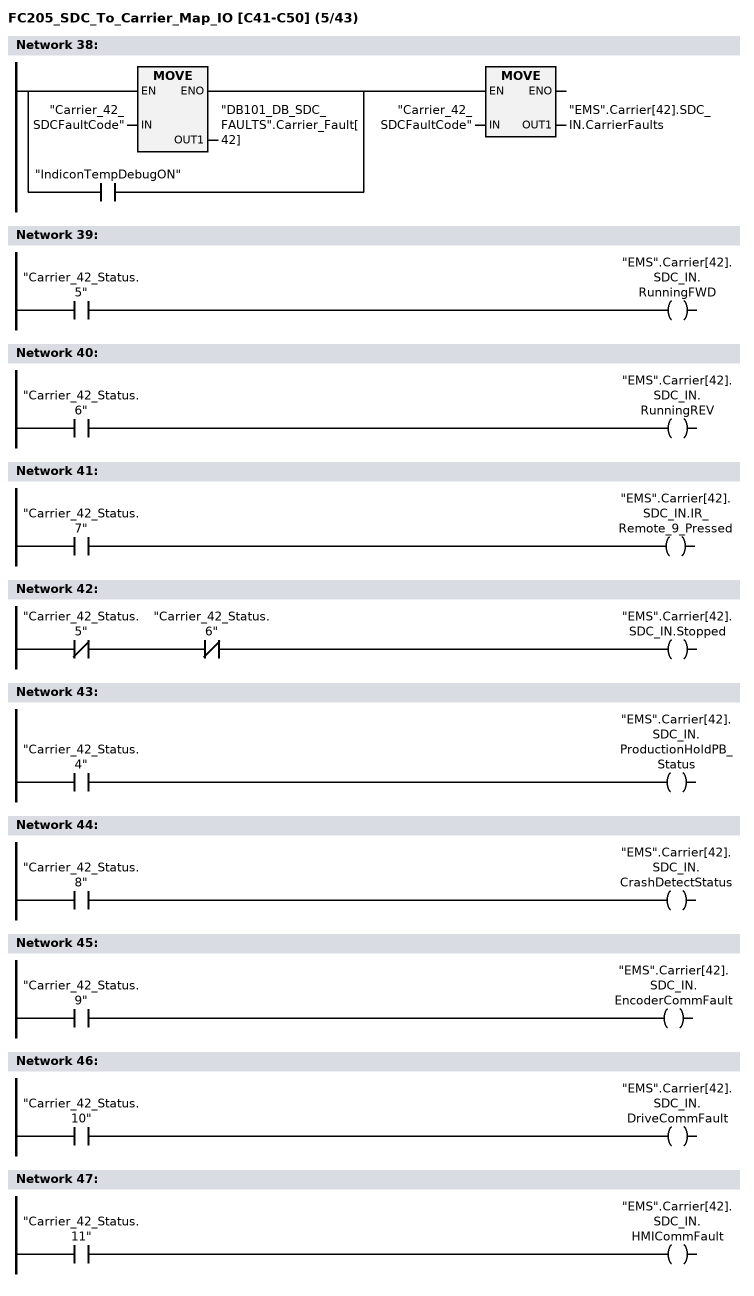
   RUNG wire#powerrail
      Move(in := "Carrier_42_SDCFaultCode", out1 => "DB101_DB_SDC_FAULTS".Carrier_Fault[42])
      wire#w1
      Move(in := "Carrier_42_SDCFaultCode", out1 => "EMS".Carrier[42].SDC_IN.CarrierFaults)
   END_RUNG
   RUNG wire#powerrail
      Contact( "IndiconTempDebugON" )
   END_RUNG wire#w1
   // the same network as SCL:
   "DB101_DB_SDC_FAULTS".Carrier_Fault[42] := "Carrier_42_SDCFaultCode";
   IF TRUE OR "IndiconTempDebugON" THEN
       "EMS".Carrier[42].SDC_IN.CarrierFaults := "Carrier_42_SDCFaultCode";
   END_IF;
END_REGION

REGION Network 39
   RUNG wire#powerrail
      Contact( "Carrier_42_Status.5" )
      Coil( "EMS".Carrier[42].SDC_IN.RunningFWD )
   END_RUNG
   // the same network as SCL:
   "EMS".Carrier[42].SDC_IN.RunningFWD := "Carrier_42_Status.5";
END_REGION

REGION Network 40
   RUNG wire#powerrail
      Contact( "Carrier_42_Status.6" )
      Coil( "EMS".Carrier[42].SDC_IN.RunningREV )
   END_RUNG
   // the same network as SCL:
   "EMS".Carrier[42].SDC_IN.RunningREV := "Carrier_42_Status.6";
END_REGION

REGION Network 41
   RUNG wire#powerrail
      Contact( "Carrier_42_Status.7" )
      Coil( "EMS".Carrier[42].SDC_IN.IR_Remote_9_Pressed )
   END_RUNG
   // the same network as SCL:
   "EMS".Carrier[42].SDC_IN.IR_Remote_9_Pressed := "Carrier_42_Status.7";
END_REGION

REGION Network 42
   RUNG wire#powerrail
      I_Contact( "Carrier_42_Status.5" )
      I_Contact( "Carrier_42_Status.6" )
      Coil( "EMS".Carrier[42].SDC_IN.Stopped )
   END_RUNG
   // the same network as SCL:
   "EMS".Carrier[42].SDC_IN.Stopped := NOT "Carrier_42_Status.5" AND NOT "Carrier_42_Status.6";
END_REGION

REGION Network 43
   RUNG wire#powerrail
      Contact( "Carrier_42_Status.4" )
      Coil( "EMS".Carrier[42].SDC_IN.ProductionHoldPB_Status )
   END_RUNG
   // the same network as SCL:
   "EMS".Carrier[42].SDC_IN.ProductionHoldPB_Status := "Carrier_42_Status.4";
END_REGION

REGION Network 44
   RUNG wire#powerrail
      Contact( "Carrier_42_Status.8" )
      Coil( "EMS".Carrier[42].SDC_IN.CrashDetectStatus )
   END_RUNG
   // the same network as SCL:
   "EMS".Carrier[42].SDC_IN.CrashDetectStatus := "Carrier_42_Status.8";
END_REGION

REGION Network 45
   RUNG wire#powerrail
      Contact( "Carrier_42_Status.9" )
      Coil( "EMS".Carrier[42].SDC_IN.EncoderCommFault )
   END_RUNG
   // the same network as SCL:
   "EMS".Carrier[42].SDC_IN.EncoderCommFault := "Carrier_42_Status.9";
END_REGION

REGION Network 46
   RUNG wire#powerrail
      Contact( "Carrier_42_Status.10" )
      Coil( "EMS".Carrier[42].SDC_IN.DriveCommFault )
   END_RUNG
   // the same network as SCL:
   "EMS".Carrier[42].SDC_IN.DriveCommFault := "Carrier_42_Status.10";
END_REGION

REGION Network 47
   RUNG wire#powerrail
      Contact( "Carrier_42_Status.11" )
      Coil( "EMS".Carrier[42].SDC_IN.HMICommFault )
   END_RUNG
   // the same network as SCL:
   "EMS".Carrier[42].SDC_IN.HMICommFault := "Carrier_42_Status.11";
END_REGION

REGION Network 48
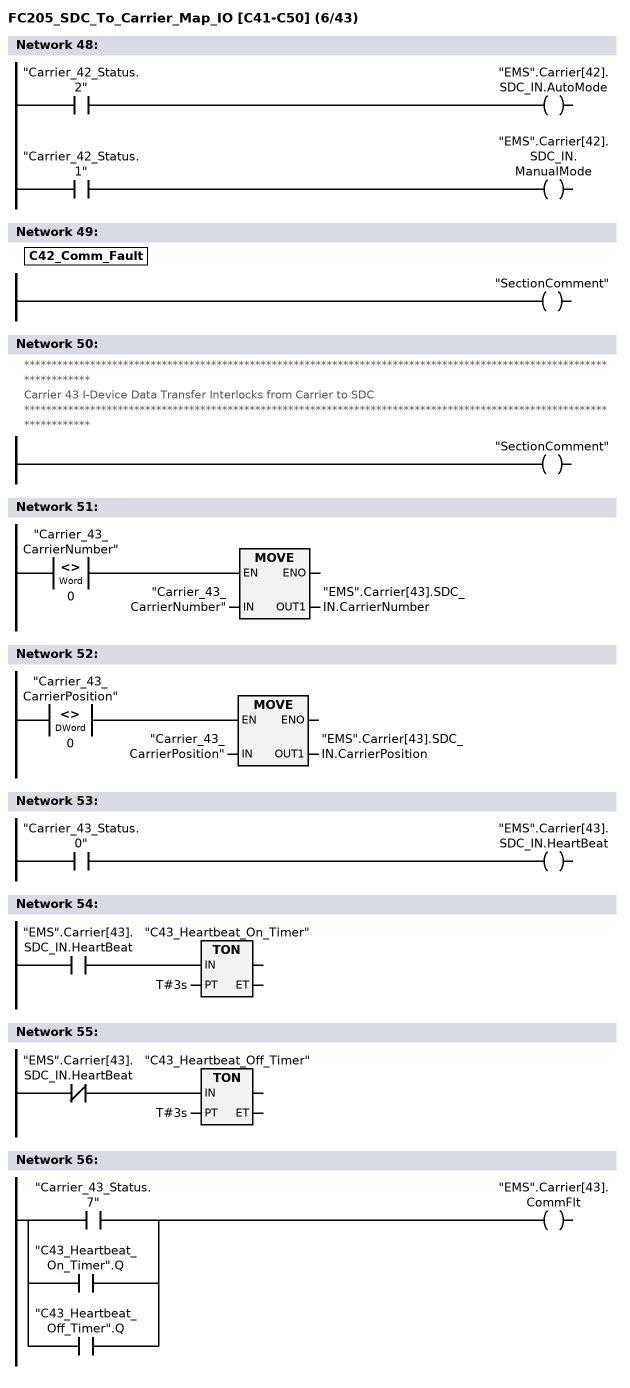
   RUNG wire#powerrail
      Contact( "Carrier_42_Status.2" )
      Coil( "EMS".Carrier[42].SDC_IN.AutoMode )
   END_RUNG
   RUNG wire#powerrail
      Contact( "Carrier_42_Status.1" )
      Coil( "EMS".Carrier[42].SDC_IN.ManualMode )
   END_RUNG
   // the same network as SCL:
   "EMS".Carrier[42].SDC_IN.AutoMode := "Carrier_42_Status.2";
   "EMS".Carrier[42].SDC_IN.ManualMode := "Carrier_42_Status.1";
END_REGION

REGION Network 49
   Label( C42_Comm_Fault )
   RUNG wire#powerrail
      Coil( "SectionComment" )
   END_RUNG
   // the same network as SCL:
   C42_Comm_Fault:
   "SectionComment" := TRUE;
END_REGION

REGION Network 50
   // **********************************************************************************************************************
   // 
   // Carrier 43 I-Device Data Transfer Interlocks from Carrier to SDC
   // 
   // **********************************************************************************************************************
   RUNG wire#powerrail
      Coil( "SectionComment" )
   END_RUNG
   // the same network as SCL:
   "SectionComment" := TRUE;
END_REGION

REGION Network 51
   RUNG wire#powerrail
      { S7_Templates := "SrcType := Word" } NE_Contact(in1 := "Carrier_43_CarrierNumber", in2 := 0)
      Move(in := "Carrier_43_CarrierNumber", out1 => "EMS".Carrier[43].SDC_IN.CarrierNumber)
   END_RUNG
   // the same network as SCL:
   IF "Carrier_43_CarrierNumber" <> 0 THEN
       "EMS".Carrier[43].SDC_IN.CarrierNumber := "Carrier_43_CarrierNumber";
   END_IF;
END_REGION

REGION Network 52
   RUNG wire#powerrail
      { S7_Templates := "SrcType := DWord" } NE_Contact(in1 := "Carrier_43_CarrierPosition", in2 := 0)
      Move(in := "Carrier_43_CarrierPosition", out1 => "EMS".Carrier[43].SDC_IN.CarrierPosition)
   END_RUNG
   // the same network as SCL:
   IF "Carrier_43_CarrierPosition" <> 0 THEN
       "EMS".Carrier[43].SDC_IN.CarrierPosition := "Carrier_43_CarrierPosition";
   END_IF;
END_REGION

REGION Network 53
   RUNG wire#powerrail
      Contact( "Carrier_43_Status.0" )
      Coil( "EMS".Carrier[43].SDC_IN.HeartBeat )
   END_RUNG
   // the same network as SCL:
   "EMS".Carrier[43].SDC_IN.HeartBeat := "Carrier_43_Status.0";
END_REGION

REGION Network 54
   "C43_Heartbeat_On_Timer".TON(IN := "EMS".Carrier[43].SDC_IN.HeartBeat, PT := T#3s);
END_REGION

REGION Network 55
   "C43_Heartbeat_Off_Timer".TON(IN := NOT "EMS".Carrier[43].SDC_IN.HeartBeat, PT := T#3s);
END_REGION

REGION Network 56
   RUNG wire#powerrail
      Contact( "Carrier_43_Status.7" )
      wire#w1
      Coil( "EMS".Carrier[43].CommFlt )
   END_RUNG
   RUNG wire#powerrail
      Contact( "C43_Heartbeat_On_Timer".Q )
   END_RUNG wire#w1
   RUNG wire#powerrail
      Contact( "C43_Heartbeat_Off_Timer".Q )
   END_RUNG wire#w1
   // the same network as SCL:
   "EMS".Carrier[43].CommFlt := "Carrier_43_Status.7" OR "C43_Heartbeat_On_Timer".Q OR "C43_Heartbeat_Off_Timer".Q;
END_REGION

REGION Network 57
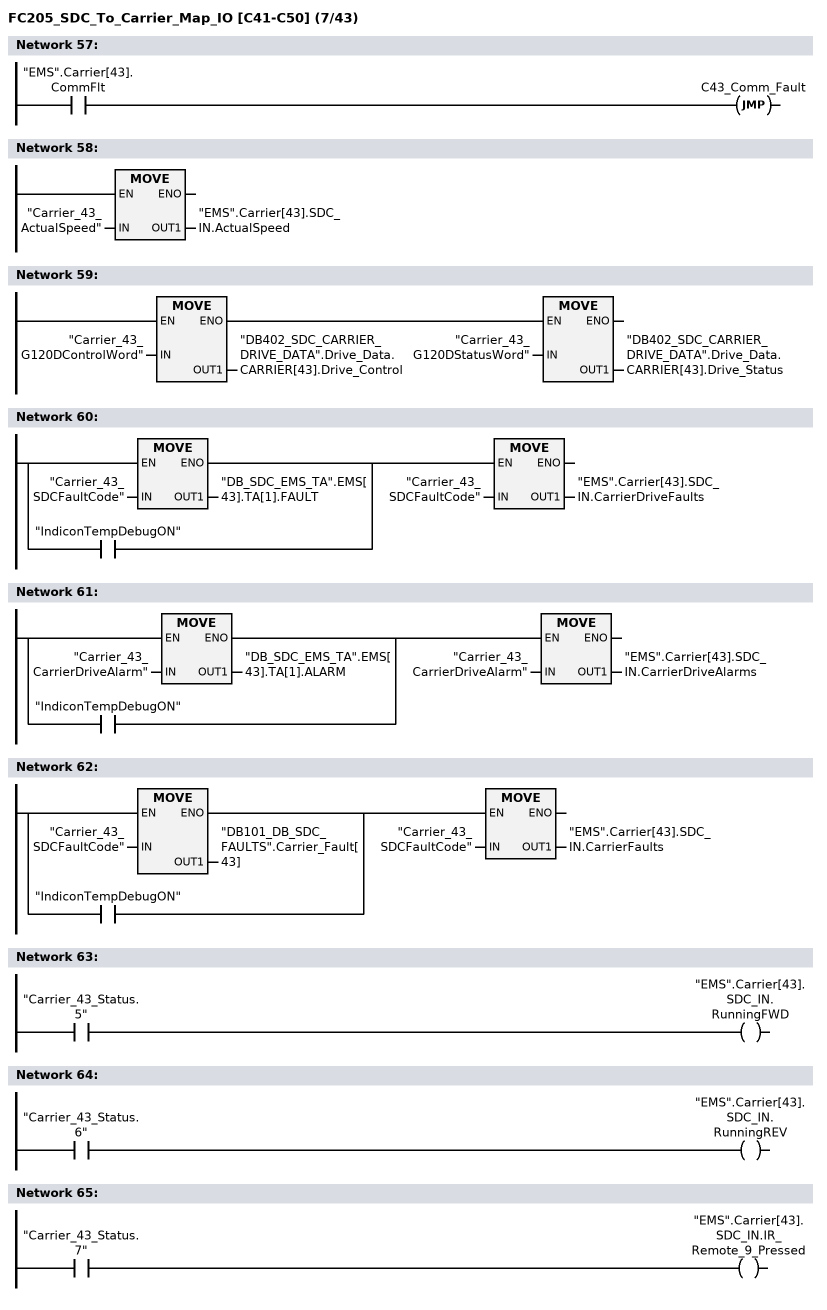
   RUNG wire#powerrail
      Contact( "EMS".Carrier[43].CommFlt )
      JumpCoil( C43_Comm_Fault )
   END_RUNG
   // the same network as SCL:
   IF "EMS".Carrier[43].CommFlt THEN GOTO C43_Comm_Fault; END_IF;
END_REGION

REGION Network 58
   RUNG wire#powerrail
      Move(in := "Carrier_43_ActualSpeed", out1 => "EMS".Carrier[43].SDC_IN.ActualSpeed)
   END_RUNG
   // the same network as SCL:
   "EMS".Carrier[43].SDC_IN.ActualSpeed := "Carrier_43_ActualSpeed";
END_REGION

REGION Network 59
   RUNG wire#powerrail
      Move(in := "Carrier_43_G120DControlWord", out1 => "DB402_SDC_CARRIER_DRIVE_DATA".Drive_Data.CARRIER[43].Drive_Control)
      Move(in := "Carrier_43_G120DStatusWord", out1 => "DB402_SDC_CARRIER_DRIVE_DATA".Drive_Data.CARRIER[43].Drive_Status)
   END_RUNG
   // the same network as SCL:
   "DB402_SDC_CARRIER_DRIVE_DATA".Drive_Data.CARRIER[43].Drive_Control := "Carrier_43_G120DControlWord";
   "DB402_SDC_CARRIER_DRIVE_DATA".Drive_Data.CARRIER[43].Drive_Status := "Carrier_43_G120DStatusWord";
END_REGION

REGION Network 60
   RUNG wire#powerrail
      Move(in := "Carrier_43_SDCFaultCode", out1 => "DB_SDC_EMS_TA".EMS[43].TA[1].FAULT)
      wire#w1
      Move(in := "Carrier_43_SDCFaultCode", out1 => "EMS".Carrier[43].SDC_IN.CarrierDriveFaults)
   END_RUNG
   RUNG wire#powerrail
      Contact( "IndiconTempDebugON" )
   END_RUNG wire#w1
   // the same network as SCL:
   "DB_SDC_EMS_TA".EMS[43].TA[1].FAULT := "Carrier_43_SDCFaultCode";
   IF TRUE OR "IndiconTempDebugON" THEN
       "EMS".Carrier[43].SDC_IN.CarrierDriveFaults := "Carrier_43_SDCFaultCode";
   END_IF;
END_REGION

REGION Network 61
   RUNG wire#powerrail
      Move(in := "Carrier_43_CarrierDriveAlarm", out1 => "DB_SDC_EMS_TA".EMS[43].TA[1].ALARM)
      wire#w1
      Move(in := "Carrier_43_CarrierDriveAlarm", out1 => "EMS".Carrier[43].SDC_IN.CarrierDriveAlarms)
   END_RUNG
   RUNG wire#powerrail
      Contact( "IndiconTempDebugON" )
   END_RUNG wire#w1
   // the same network as SCL:
   "DB_SDC_EMS_TA".EMS[43].TA[1].ALARM := "Carrier_43_CarrierDriveAlarm";
   IF TRUE OR "IndiconTempDebugON" THEN
       "EMS".Carrier[43].SDC_IN.CarrierDriveAlarms := "Carrier_43_CarrierDriveAlarm";
   END_IF;
END_REGION

REGION Network 62
   RUNG wire#powerrail
      Move(in := "Carrier_43_SDCFaultCode", out1 => "DB101_DB_SDC_FAULTS".Carrier_Fault[43])
      wire#w1
      Move(in := "Carrier_43_SDCFaultCode", out1 => "EMS".Carrier[43].SDC_IN.CarrierFaults)
   END_RUNG
   RUNG wire#powerrail
      Contact( "IndiconTempDebugON" )
   END_RUNG wire#w1
   // the same network as SCL:
   "DB101_DB_SDC_FAULTS".Carrier_Fault[43] := "Carrier_43_SDCFaultCode";
   IF TRUE OR "IndiconTempDebugON" THEN
       "EMS".Carrier[43].SDC_IN.CarrierFaults := "Carrier_43_SDCFaultCode";
   END_IF;
END_REGION

REGION Network 63
   RUNG wire#powerrail
      Contact( "Carrier_43_Status.5" )
      Coil( "EMS".Carrier[43].SDC_IN.RunningFWD )
   END_RUNG
   // the same network as SCL:
   "EMS".Carrier[43].SDC_IN.RunningFWD := "Carrier_43_Status.5";
END_REGION

REGION Network 64
   RUNG wire#powerrail
      Contact( "Carrier_43_Status.6" )
      Coil( "EMS".Carrier[43].SDC_IN.RunningREV )
   END_RUNG
   // the same network as SCL:
   "EMS".Carrier[43].SDC_IN.RunningREV := "Carrier_43_Status.6";
END_REGION

REGION Network 65
   RUNG wire#powerrail
      Contact( "Carrier_43_Status.7" )
      Coil( "EMS".Carrier[43].SDC_IN.IR_Remote_9_Pressed )
   END_RUNG
   // the same network as SCL:
   "EMS".Carrier[43].SDC_IN.IR_Remote_9_Pressed := "Carrier_43_Status.7";
END_REGION

REGION Network 66
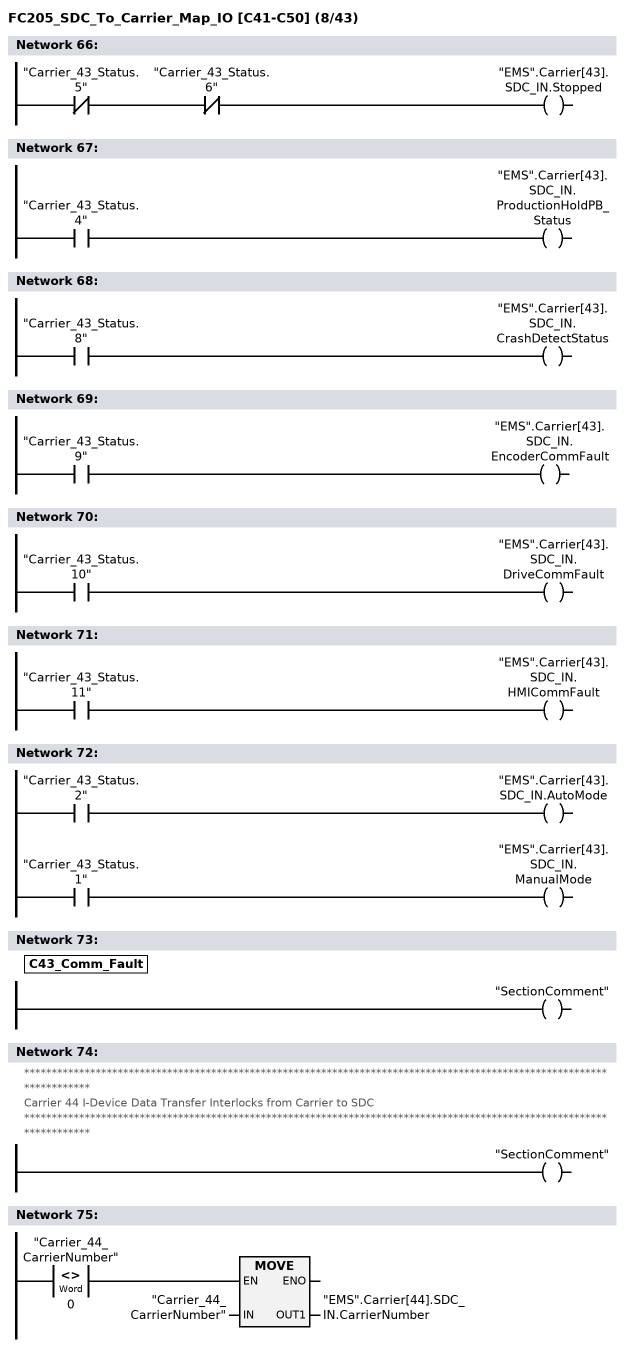
   RUNG wire#powerrail
      I_Contact( "Carrier_43_Status.5" )
      I_Contact( "Carrier_43_Status.6" )
      Coil( "EMS".Carrier[43].SDC_IN.Stopped )
   END_RUNG
   // the same network as SCL:
   "EMS".Carrier[43].SDC_IN.Stopped := NOT "Carrier_43_Status.5" AND NOT "Carrier_43_Status.6";
END_REGION

REGION Network 67
   RUNG wire#powerrail
      Contact( "Carrier_43_Status.4" )
      Coil( "EMS".Carrier[43].SDC_IN.ProductionHoldPB_Status )
   END_RUNG
   // the same network as SCL:
   "EMS".Carrier[43].SDC_IN.ProductionHoldPB_Status := "Carrier_43_Status.4";
END_REGION

REGION Network 68
   RUNG wire#powerrail
      Contact( "Carrier_43_Status.8" )
      Coil( "EMS".Carrier[43].SDC_IN.CrashDetectStatus )
   END_RUNG
   // the same network as SCL:
   "EMS".Carrier[43].SDC_IN.CrashDetectStatus := "Carrier_43_Status.8";
END_REGION

REGION Network 69
   RUNG wire#powerrail
      Contact( "Carrier_43_Status.9" )
      Coil( "EMS".Carrier[43].SDC_IN.EncoderCommFault )
   END_RUNG
   // the same network as SCL:
   "EMS".Carrier[43].SDC_IN.EncoderCommFault := "Carrier_43_Status.9";
END_REGION

REGION Network 70
   RUNG wire#powerrail
      Contact( "Carrier_43_Status.10" )
      Coil( "EMS".Carrier[43].SDC_IN.DriveCommFault )
   END_RUNG
   // the same network as SCL:
   "EMS".Carrier[43].SDC_IN.DriveCommFault := "Carrier_43_Status.10";
END_REGION

REGION Network 71
   RUNG wire#powerrail
      Contact( "Carrier_43_Status.11" )
      Coil( "EMS".Carrier[43].SDC_IN.HMICommFault )
   END_RUNG
   // the same network as SCL:
   "EMS".Carrier[43].SDC_IN.HMICommFault := "Carrier_43_Status.11";
END_REGION

REGION Network 72
   RUNG wire#powerrail
      Contact( "Carrier_43_Status.2" )
      Coil( "EMS".Carrier[43].SDC_IN.AutoMode )
   END_RUNG
   RUNG wire#powerrail
      Contact( "Carrier_43_Status.1" )
      Coil( "EMS".Carrier[43].SDC_IN.ManualMode )
   END_RUNG
   // the same network as SCL:
   "EMS".Carrier[43].SDC_IN.AutoMode := "Carrier_43_Status.2";
   "EMS".Carrier[43].SDC_IN.ManualMode := "Carrier_43_Status.1";
END_REGION

REGION Network 73
   Label( C43_Comm_Fault )
   RUNG wire#powerrail
      Coil( "SectionComment" )
   END_RUNG
   // the same network as SCL:
   C43_Comm_Fault:
   "SectionComment" := TRUE;
END_REGION

REGION Network 74
   // **********************************************************************************************************************
   // 
   // Carrier 44 I-Device Data Transfer Interlocks from Carrier to SDC
   // 
   // **********************************************************************************************************************
   RUNG wire#powerrail
      Coil( "SectionComment" )
   END_RUNG
   // the same network as SCL:
   "SectionComment" := TRUE;
END_REGION

REGION Network 75
   RUNG wire#powerrail
      { S7_Templates := "SrcType := Word" } NE_Contact(in1 := "Carrier_44_CarrierNumber", in2 := 0)
      Move(in := "Carrier_44_CarrierNumber", out1 => "EMS".Carrier[44].SDC_IN.CarrierNumber)
   END_RUNG
   // the same network as SCL:
   IF "Carrier_44_CarrierNumber" <> 0 THEN
       "EMS".Carrier[44].SDC_IN.CarrierNumber := "Carrier_44_CarrierNumber";
   END_IF;
END_REGION

REGION Network 76
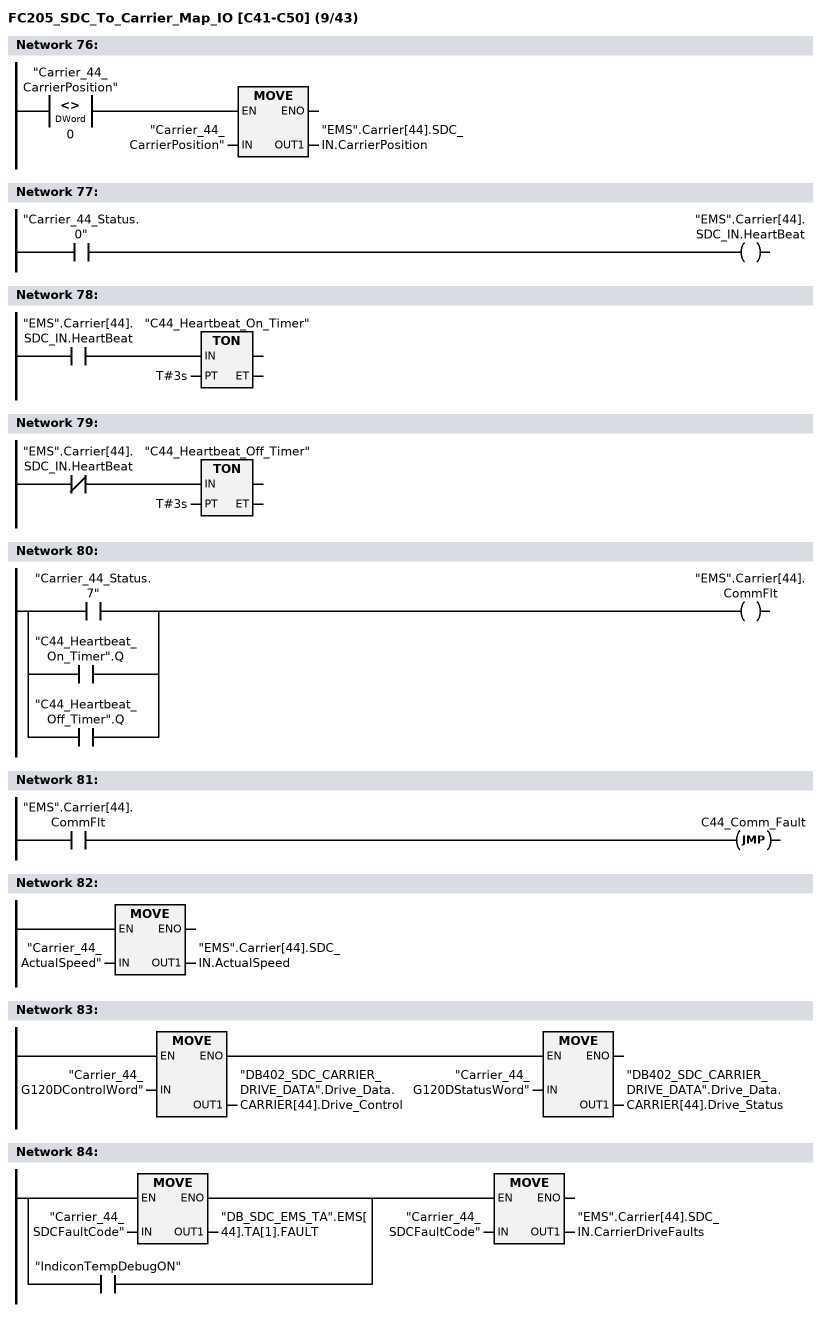
   RUNG wire#powerrail
      { S7_Templates := "SrcType := DWord" } NE_Contact(in1 := "Carrier_44_CarrierPosition", in2 := 0)
      Move(in := "Carrier_44_CarrierPosition", out1 => "EMS".Carrier[44].SDC_IN.CarrierPosition)
   END_RUNG
   // the same network as SCL:
   IF "Carrier_44_CarrierPosition" <> 0 THEN
       "EMS".Carrier[44].SDC_IN.CarrierPosition := "Carrier_44_CarrierPosition";
   END_IF;
END_REGION

REGION Network 77
   RUNG wire#powerrail
      Contact( "Carrier_44_Status.0" )
      Coil( "EMS".Carrier[44].SDC_IN.HeartBeat )
   END_RUNG
   // the same network as SCL:
   "EMS".Carrier[44].SDC_IN.HeartBeat := "Carrier_44_Status.0";
END_REGION

REGION Network 78
   "C44_Heartbeat_On_Timer".TON(IN := "EMS".Carrier[44].SDC_IN.HeartBeat, PT := T#3s);
END_REGION

REGION Network 79
   "C44_Heartbeat_Off_Timer".TON(IN := NOT "EMS".Carrier[44].SDC_IN.HeartBeat, PT := T#3s);
END_REGION

REGION Network 80
   RUNG wire#powerrail
      Contact( "Carrier_44_Status.7" )
      wire#w1
      Coil( "EMS".Carrier[44].CommFlt )
   END_RUNG
   RUNG wire#powerrail
      Contact( "C44_Heartbeat_On_Timer".Q )
   END_RUNG wire#w1
   RUNG wire#powerrail
      Contact( "C44_Heartbeat_Off_Timer".Q )
   END_RUNG wire#w1
   // the same network as SCL:
   "EMS".Carrier[44].CommFlt := "Carrier_44_Status.7" OR "C44_Heartbeat_On_Timer".Q OR "C44_Heartbeat_Off_Timer".Q;
END_REGION

REGION Network 81
   RUNG wire#powerrail
      Contact( "EMS".Carrier[44].CommFlt )
      JumpCoil( C44_Comm_Fault )
   END_RUNG
   // the same network as SCL:
   IF "EMS".Carrier[44].CommFlt THEN GOTO C44_Comm_Fault; END_IF;
END_REGION

REGION Network 82
   RUNG wire#powerrail
      Move(in := "Carrier_44_ActualSpeed", out1 => "EMS".Carrier[44].SDC_IN.ActualSpeed)
   END_RUNG
   // the same network as SCL:
   "EMS".Carrier[44].SDC_IN.ActualSpeed := "Carrier_44_ActualSpeed";
END_REGION

REGION Network 83
   RUNG wire#powerrail
      Move(in := "Carrier_44_G120DControlWord", out1 => "DB402_SDC_CARRIER_DRIVE_DATA".Drive_Data.CARRIER[44].Drive_Control)
      Move(in := "Carrier_44_G120DStatusWord", out1 => "DB402_SDC_CARRIER_DRIVE_DATA".Drive_Data.CARRIER[44].Drive_Status)
   END_RUNG
   // the same network as SCL:
   "DB402_SDC_CARRIER_DRIVE_DATA".Drive_Data.CARRIER[44].Drive_Control := "Carrier_44_G120DControlWord";
   "DB402_SDC_CARRIER_DRIVE_DATA".Drive_Data.CARRIER[44].Drive_Status := "Carrier_44_G120DStatusWord";
END_REGION

REGION Network 84
   RUNG wire#powerrail
      Move(in := "Carrier_44_SDCFaultCode", out1 => "DB_SDC_EMS_TA".EMS[44].TA[1].FAULT)
      wire#w1
      Move(in := "Carrier_44_SDCFaultCode", out1 => "EMS".Carrier[44].SDC_IN.CarrierDriveFaults)
   END_RUNG
   RUNG wire#powerrail
      Contact( "IndiconTempDebugON" )
   END_RUNG wire#w1
   // the same network as SCL:
   "DB_SDC_EMS_TA".EMS[44].TA[1].FAULT := "Carrier_44_SDCFaultCode";
   IF TRUE OR "IndiconTempDebugON" THEN
       "EMS".Carrier[44].SDC_IN.CarrierDriveFaults := "Carrier_44_SDCFaultCode";
   END_IF;
END_REGION

REGION Network 85
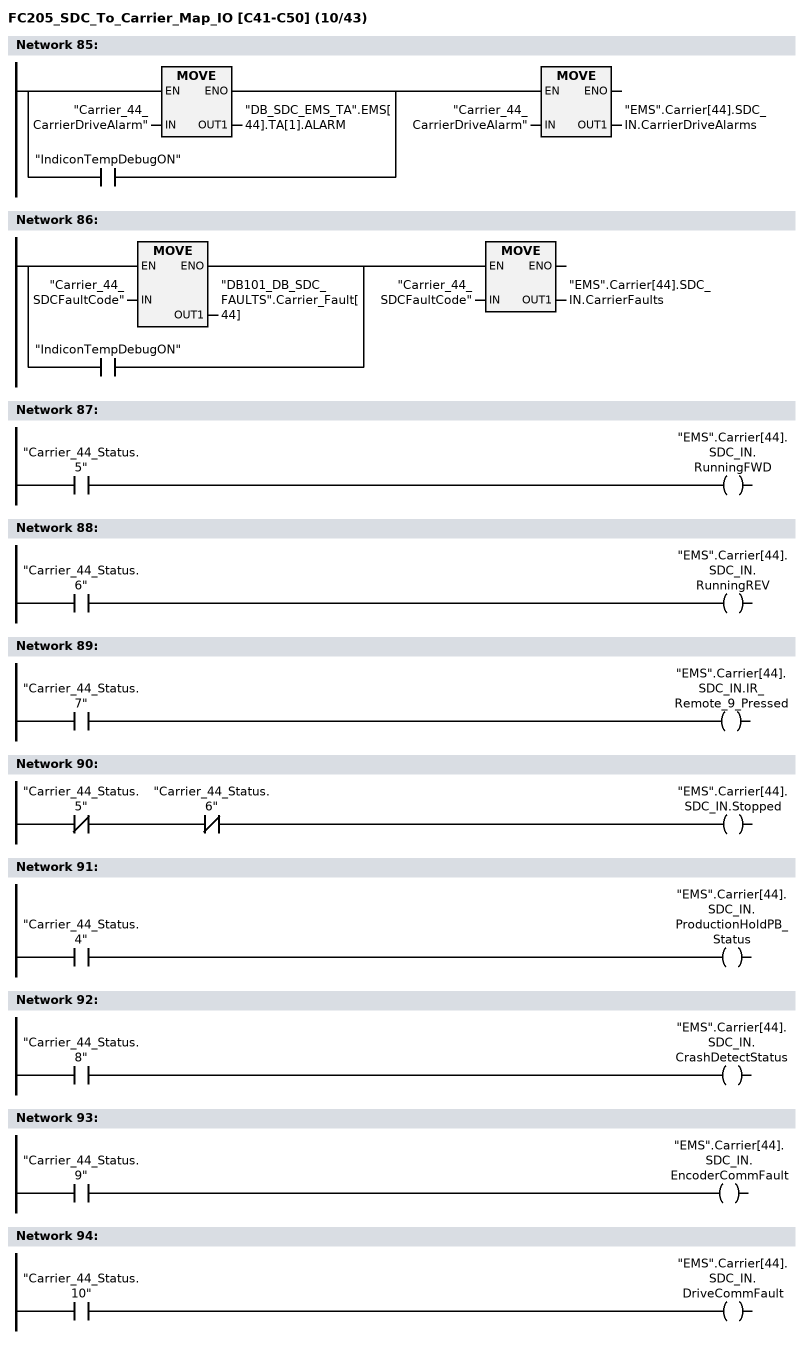
   RUNG wire#powerrail
      Move(in := "Carrier_44_CarrierDriveAlarm", out1 => "DB_SDC_EMS_TA".EMS[44].TA[1].ALARM)
      wire#w1
      Move(in := "Carrier_44_CarrierDriveAlarm", out1 => "EMS".Carrier[44].SDC_IN.CarrierDriveAlarms)
   END_RUNG
   RUNG wire#powerrail
      Contact( "IndiconTempDebugON" )
   END_RUNG wire#w1
   // the same network as SCL:
   "DB_SDC_EMS_TA".EMS[44].TA[1].ALARM := "Carrier_44_CarrierDriveAlarm";
   IF TRUE OR "IndiconTempDebugON" THEN
       "EMS".Carrier[44].SDC_IN.CarrierDriveAlarms := "Carrier_44_CarrierDriveAlarm";
   END_IF;
END_REGION

REGION Network 86
   RUNG wire#powerrail
      Move(in := "Carrier_44_SDCFaultCode", out1 => "DB101_DB_SDC_FAULTS".Carrier_Fault[44])
      wire#w1
      Move(in := "Carrier_44_SDCFaultCode", out1 => "EMS".Carrier[44].SDC_IN.CarrierFaults)
   END_RUNG
   RUNG wire#powerrail
      Contact( "IndiconTempDebugON" )
   END_RUNG wire#w1
   // the same network as SCL:
   "DB101_DB_SDC_FAULTS".Carrier_Fault[44] := "Carrier_44_SDCFaultCode";
   IF TRUE OR "IndiconTempDebugON" THEN
       "EMS".Carrier[44].SDC_IN.CarrierFaults := "Carrier_44_SDCFaultCode";
   END_IF;
END_REGION

REGION Network 87
   RUNG wire#powerrail
      Contact( "Carrier_44_Status.5" )
      Coil( "EMS".Carrier[44].SDC_IN.RunningFWD )
   END_RUNG
   // the same network as SCL:
   "EMS".Carrier[44].SDC_IN.RunningFWD := "Carrier_44_Status.5";
END_REGION

REGION Network 88
   RUNG wire#powerrail
      Contact( "Carrier_44_Status.6" )
      Coil( "EMS".Carrier[44].SDC_IN.RunningREV )
   END_RUNG
   // the same network as SCL:
   "EMS".Carrier[44].SDC_IN.RunningREV := "Carrier_44_Status.6";
END_REGION

REGION Network 89
   RUNG wire#powerrail
      Contact( "Carrier_44_Status.7" )
      Coil( "EMS".Carrier[44].SDC_IN.IR_Remote_9_Pressed )
   END_RUNG
   // the same network as SCL:
   "EMS".Carrier[44].SDC_IN.IR_Remote_9_Pressed := "Carrier_44_Status.7";
END_REGION

REGION Network 90
   RUNG wire#powerrail
      I_Contact( "Carrier_44_Status.5" )
      I_Contact( "Carrier_44_Status.6" )
      Coil( "EMS".Carrier[44].SDC_IN.Stopped )
   END_RUNG
   // the same network as SCL:
   "EMS".Carrier[44].SDC_IN.Stopped := NOT "Carrier_44_Status.5" AND NOT "Carrier_44_Status.6";
END_REGION

REGION Network 91
   RUNG wire#powerrail
      Contact( "Carrier_44_Status.4" )
      Coil( "EMS".Carrier[44].SDC_IN.ProductionHoldPB_Status )
   END_RUNG
   // the same network as SCL:
   "EMS".Carrier[44].SDC_IN.ProductionHoldPB_Status := "Carrier_44_Status.4";
END_REGION

REGION Network 92
   RUNG wire#powerrail
      Contact( "Carrier_44_Status.8" )
      Coil( "EMS".Carrier[44].SDC_IN.CrashDetectStatus )
   END_RUNG
   // the same network as SCL:
   "EMS".Carrier[44].SDC_IN.CrashDetectStatus := "Carrier_44_Status.8";
END_REGION

REGION Network 93
   RUNG wire#powerrail
      Contact( "Carrier_44_Status.9" )
      Coil( "EMS".Carrier[44].SDC_IN.EncoderCommFault )
   END_RUNG
   // the same network as SCL:
   "EMS".Carrier[44].SDC_IN.EncoderCommFault := "Carrier_44_Status.9";
END_REGION

REGION Network 94
   RUNG wire#powerrail
      Contact( "Carrier_44_Status.10" )
      Coil( "EMS".Carrier[44].SDC_IN.DriveCommFault )
   END_RUNG
   // the same network as SCL:
   "EMS".Carrier[44].SDC_IN.DriveCommFault := "Carrier_44_Status.10";
END_REGION

REGION Network 95
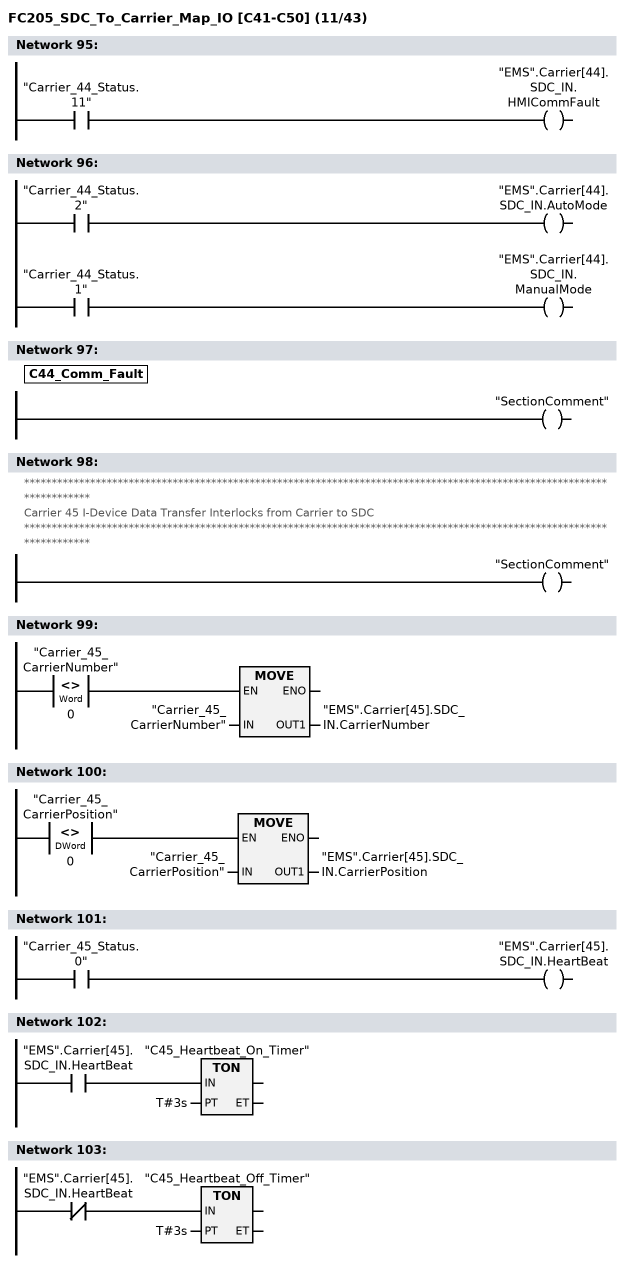
   RUNG wire#powerrail
      Contact( "Carrier_44_Status.11" )
      Coil( "EMS".Carrier[44].SDC_IN.HMICommFault )
   END_RUNG
   // the same network as SCL:
   "EMS".Carrier[44].SDC_IN.HMICommFault := "Carrier_44_Status.11";
END_REGION

REGION Network 96
   RUNG wire#powerrail
      Contact( "Carrier_44_Status.2" )
      Coil( "EMS".Carrier[44].SDC_IN.AutoMode )
   END_RUNG
   RUNG wire#powerrail
      Contact( "Carrier_44_Status.1" )
      Coil( "EMS".Carrier[44].SDC_IN.ManualMode )
   END_RUNG
   // the same network as SCL:
   "EMS".Carrier[44].SDC_IN.AutoMode := "Carrier_44_Status.2";
   "EMS".Carrier[44].SDC_IN.ManualMode := "Carrier_44_Status.1";
END_REGION

REGION Network 97
   Label( C44_Comm_Fault )
   RUNG wire#powerrail
      Coil( "SectionComment" )
   END_RUNG
   // the same network as SCL:
   C44_Comm_Fault:
   "SectionComment" := TRUE;
END_REGION

REGION Network 98
   // **********************************************************************************************************************
   // 
   // Carrier 45 I-Device Data Transfer Interlocks from Carrier to SDC
   // 
   // **********************************************************************************************************************
   RUNG wire#powerrail
      Coil( "SectionComment" )
   END_RUNG
   // the same network as SCL:
   "SectionComment" := TRUE;
END_REGION

REGION Network 99
   RUNG wire#powerrail
      { S7_Templates := "SrcType := Word" } NE_Contact(in1 := "Carrier_45_CarrierNumber", in2 := 0)
      Move(in := "Carrier_45_CarrierNumber", out1 => "EMS".Carrier[45].SDC_IN.CarrierNumber)
   END_RUNG
   // the same network as SCL:
   IF "Carrier_45_CarrierNumber" <> 0 THEN
       "EMS".Carrier[45].SDC_IN.CarrierNumber := "Carrier_45_CarrierNumber";
   END_IF;
END_REGION

REGION Network 100
   RUNG wire#powerrail
      { S7_Templates := "SrcType := DWord" } NE_Contact(in1 := "Carrier_45_CarrierPosition", in2 := 0)
      Move(in := "Carrier_45_CarrierPosition", out1 => "EMS".Carrier[45].SDC_IN.CarrierPosition)
   END_RUNG
   // the same network as SCL:
   IF "Carrier_45_CarrierPosition" <> 0 THEN
       "EMS".Carrier[45].SDC_IN.CarrierPosition := "Carrier_45_CarrierPosition";
   END_IF;
END_REGION

REGION Network 101
   RUNG wire#powerrail
      Contact( "Carrier_45_Status.0" )
      Coil( "EMS".Carrier[45].SDC_IN.HeartBeat )
   END_RUNG
   // the same network as SCL:
   "EMS".Carrier[45].SDC_IN.HeartBeat := "Carrier_45_Status.0";
END_REGION

REGION Network 102
   "C45_Heartbeat_On_Timer".TON(IN := "EMS".Carrier[45].SDC_IN.HeartBeat, PT := T#3s);
END_REGION

REGION Network 103
   "C45_Heartbeat_Off_Timer".TON(IN := NOT "EMS".Carrier[45].SDC_IN.HeartBeat, PT := T#3s);
END_REGION

REGION Network 104
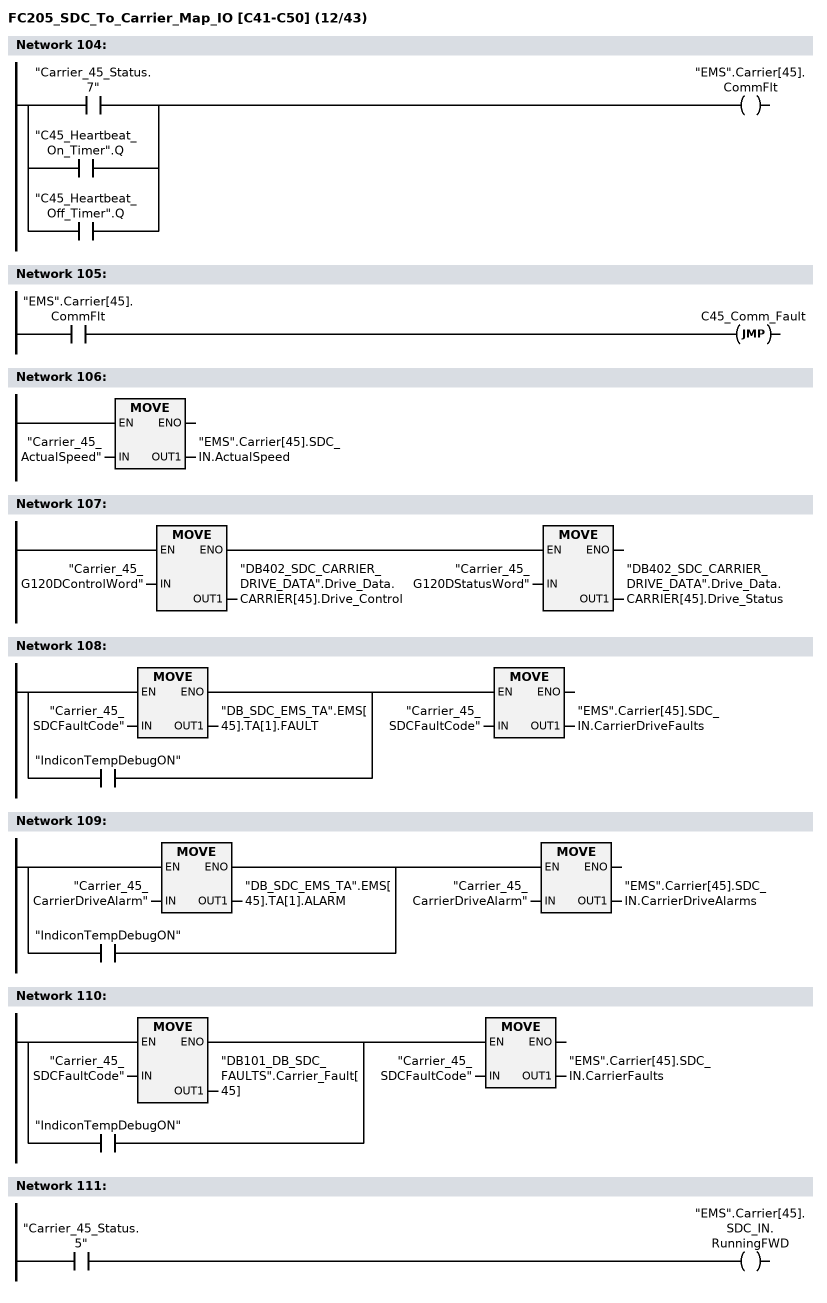
   RUNG wire#powerrail
      Contact( "Carrier_45_Status.7" )
      wire#w1
      Coil( "EMS".Carrier[45].CommFlt )
   END_RUNG
   RUNG wire#powerrail
      Contact( "C45_Heartbeat_On_Timer".Q )
   END_RUNG wire#w1
   RUNG wire#powerrail
      Contact( "C45_Heartbeat_Off_Timer".Q )
   END_RUNG wire#w1
   // the same network as SCL:
   "EMS".Carrier[45].CommFlt := "Carrier_45_Status.7" OR "C45_Heartbeat_On_Timer".Q OR "C45_Heartbeat_Off_Timer".Q;
END_REGION

REGION Network 105
   RUNG wire#powerrail
      Contact( "EMS".Carrier[45].CommFlt )
      JumpCoil( C45_Comm_Fault )
   END_RUNG
   // the same network as SCL:
   IF "EMS".Carrier[45].CommFlt THEN GOTO C45_Comm_Fault; END_IF;
END_REGION

REGION Network 106
   RUNG wire#powerrail
      Move(in := "Carrier_45_ActualSpeed", out1 => "EMS".Carrier[45].SDC_IN.ActualSpeed)
   END_RUNG
   // the same network as SCL:
   "EMS".Carrier[45].SDC_IN.ActualSpeed := "Carrier_45_ActualSpeed";
END_REGION

REGION Network 107
   RUNG wire#powerrail
      Move(in := "Carrier_45_G120DControlWord", out1 => "DB402_SDC_CARRIER_DRIVE_DATA".Drive_Data.CARRIER[45].Drive_Control)
      Move(in := "Carrier_45_G120DStatusWord", out1 => "DB402_SDC_CARRIER_DRIVE_DATA".Drive_Data.CARRIER[45].Drive_Status)
   END_RUNG
   // the same network as SCL:
   "DB402_SDC_CARRIER_DRIVE_DATA".Drive_Data.CARRIER[45].Drive_Control := "Carrier_45_G120DControlWord";
   "DB402_SDC_CARRIER_DRIVE_DATA".Drive_Data.CARRIER[45].Drive_Status := "Carrier_45_G120DStatusWord";
END_REGION

REGION Network 108
   RUNG wire#powerrail
      Move(in := "Carrier_45_SDCFaultCode", out1 => "DB_SDC_EMS_TA".EMS[45].TA[1].FAULT)
      wire#w1
      Move(in := "Carrier_45_SDCFaultCode", out1 => "EMS".Carrier[45].SDC_IN.CarrierDriveFaults)
   END_RUNG
   RUNG wire#powerrail
      Contact( "IndiconTempDebugON" )
   END_RUNG wire#w1
   // the same network as SCL:
   "DB_SDC_EMS_TA".EMS[45].TA[1].FAULT := "Carrier_45_SDCFaultCode";
   IF TRUE OR "IndiconTempDebugON" THEN
       "EMS".Carrier[45].SDC_IN.CarrierDriveFaults := "Carrier_45_SDCFaultCode";
   END_IF;
END_REGION

REGION Network 109
   RUNG wire#powerrail
      Move(in := "Carrier_45_CarrierDriveAlarm", out1 => "DB_SDC_EMS_TA".EMS[45].TA[1].ALARM)
      wire#w1
      Move(in := "Carrier_45_CarrierDriveAlarm", out1 => "EMS".Carrier[45].SDC_IN.CarrierDriveAlarms)
   END_RUNG
   RUNG wire#powerrail
      Contact( "IndiconTempDebugON" )
   END_RUNG wire#w1
   // the same network as SCL:
   "DB_SDC_EMS_TA".EMS[45].TA[1].ALARM := "Carrier_45_CarrierDriveAlarm";
   IF TRUE OR "IndiconTempDebugON" THEN
       "EMS".Carrier[45].SDC_IN.CarrierDriveAlarms := "Carrier_45_CarrierDriveAlarm";
   END_IF;
END_REGION
